// TIA Portal project "Label_Process" (V20)
// Label and sorter box process

(* hardware
DEVICE "S7-1200 station_1"  S7-1200 Station
   slot 0: "Rack_0"  S7-1200 Rack  Rack  V1.0
   slot 1: "PLC_1"  CPU 1212C AC/DC/Rly  6ES7 212-1BE40-0XB0  V4.6
DEVICE "HMI_1"  TP1200 Comfort
   slot 0: "HMI_1"  TP1200 Comfort  6AV2 124-0MC01-0AX0  17.0.0.0
   slot 1: "HMI_RT_1"  TP1200 Comfort  6AV2 124-0MC01-0AX0  17.0.0.0
   slot 5: "HMI_1.IE_CP_1"  PROFINET Interface  17.0.0.0
      slot 1: "PROFINET Interface_1"  PROFINET Interface
         slot 1: "Port_1"  Port
         slot 2: "Port_2"  Port
   slot 7: "HMI_1.MPI/DP_CP_1"  MPI/DP Interface  17.0.0.0
*)

// ===== PLC "PLC_1"  CPU 1212C AC/DC/Rly =====

VAR_GLOBAL   // PLC tag table "Inputs_FactoryIO"
   "Emergency_Stop" AT %I1.0 : Bool;   // Emergency stop mushroom
   "Stop_Pb" AT %I1.1 : Bool;   // Stop pushbutton
   "Start_Pb" AT %I1.2 : Bool;   // Start pushbutton
   "Pause_Signal" AT %I1.3 : Bool;   // Selector for pause process
   "Heigh_Box" AT %I1.4 : Bool;   // Sensor for heigh box
   "Position_Box" AT %I1.5 : Bool;   // Sensor of position box at the label zone
   "Unlabel_Box" AT %I1.6 : Bool;   // Unlabel box sensor
   "Thermal_Fault" AT %I1.7 : Bool;   // Thermal Fault from thermal relays
   "Clock_Byte" AT %MB10 : Byte;
   "Clock_10Hz" AT %M10.0 : Bool;
   "Clock_5Hz" AT %M10.1 : Bool;
   "Clock_2.5Hz" AT %M10.2 : Bool;
   "Clock_2Hz" AT %M10.3 : Bool;
   "Clock_1.25Hz" AT %M10.4 : Bool;
   "Clock_1Hz" AT %M10.5 : Bool;
   "Clock_0.625Hz" AT %M10.6 : Bool;
   "Clock_0.5Hz" AT %M10.7 : Bool;
   "Tag_1" AT %M8.1 : Bool;
   "Tag_2" AT %M1.1 : Bool;
END_VAR

VAR_GLOBAL   // PLC tag table "Outputs"
   "Conveyor M1" AT %Q0.0 : Bool;   // Control Conveyor Belt M1
   "Conveyor M2" AT %Q0.1 : Bool;   // Control Conveyor Belt M2
   "Conveyor M3" AT %Q0.2 : Bool;   // Control Conveyor Belt M3
   "Sorter" AT %Q0.3 : Bool;   // Activate sorter
   "Sorter_Left" AT %Q0.4 : Bool;   // Activate sorter for left position
   "Axis_Label" AT %Q0.5 : Bool;   // Axis control for labeled
END_VAR

DATA_BLOCK "DATA"   // DB1
{ S7_Optimized_Access := 'TRUE' }
VERSION : 0.1
   VAR
      varCounters : Struct
         Labeled_Boxes_Counter : Int;   // Labeled boxes counter
         Unlabel_Boxes_Counter : Int;   // Unlabel boxes counter
         CountUp_Unlabel : Bool;
         Total_Boxes : Int;
         Reset_Counters : Bool;
         Label_TimeSec : DInt;
      END_STRUCT;
      activateSorter : Struct
         M_Sorter_Left : Bool;
         M1_Activate_Sorter : Bool;
         M2_Activate_Sorter : Bool;
      END_STRUCT;
      risingEgde : Struct
         R_StartPB : Bool;   // Memory for rising edge Start button
         R_positionBox : Bool;   // Memory for rising edge position box sensor
         R_Heigh_Box : Bool;   // Memory for rising egde heigh box sensor
         R_Unlabel_Box : Bool;   // Memory for rising egde unlabel box sensor
         R_CountUP_Unlabel : Bool;
         R_Move_CountUP : Bool;
      END_STRUCT;
      generalData : Struct
         M_startStop : Bool;   // Memory for Start Stop all process
         M_pauseProcess : Bool;   // Memory for Pause all process
      END_STRUCT;
      Belts_Data : Struct
         M_Activate_M1 : Bool;   // Memory for activate Belt Conveyor M1
         M_Activate_M2 : Bool;   // Memory for activate Belt Conveyor M2
         M_Activate_M3 : Bool;   // Memory for activate Belt Conveyor M3
      END_STRUCT;
   END_VAR
BEGIN
END_DATA_BLOCK

DATA_BLOCK "HMI_Data"   // DB3
{ S7_Optimized_Access := 'TRUE' }
VERSION : 0.1
   VAR
      "Inputs from HMI" : Struct   // Inputs signals from HMI
         startSignal : Bool;   // Start all process
         stopSignal : Bool;   // Stop all process
         resetCounters : Bool;   // Reset all counters
         pauseProcess : Bool;   // Pause all process
      END_STRUCT;
      Move_Animation : Int;   // HMI box animation
      "Belt Control" : Struct   // Start signals for each belt conveyor
         Start_M1 : Bool;   // Start belt conveyor M1
         Start_M2 : Bool;   // Start belt conveyor M2
         Start_M3 : Bool;   // Start belt conveyor M3
      END_STRUCT;
      "Sorter & Axis Control" : Struct   // Controlling sorter and axis label
         activateAxis : Bool;
         activateSorter : Bool;
         activateSorterLeft : Bool;
      END_STRUCT;
      Counters : Struct
         resetCounterLabeled : Bool;
         resetCounterUnlabel : Bool;
         labelTime : DInt;
      END_STRUCT;
   END_VAR
BEGIN
END_DATA_BLOCK

DATA_BLOCK "HMI_Alarms"   // DB4
{ S7_Optimized_Access := 'FALSE' }
VERSION : 0.1
   VAR
      noTimeSet : Bool;   // Alarm indicator, no time for axis label actuator
      emergencyStopPushed : Bool;   // Alarm indicator, emergency stop pushed
      thermalFault : Bool;   // Alarm indicator, fault thermal relays
      pauseActive : Bool;   // Warning indicator, pause active
   END_VAR
BEGIN
END_DATA_BLOCK

// folder: System blocks/Program resources

DATA_BLOCK "axisTimer"   // DB2
{ S7_Optimized_Access := 'TRUE' }
AUTHOR : Simatic
FAMILY : IEC
NAME : IEC_TMR
VERSION : 1.0
// stored: InstanceOfName IEC_TIMER
"IEC_TIMER"
BEGIN
END_DATA_BLOCK

// folder: (top level)

FUNCTION "Start_Stop" : Void   // FC1, LAD
TITLE = Start and Stop Block
{ S7_Optimized_Access := 'TRUE' }
AUTHOR : Stiven Perez
VERSION : 0.1
// Start and stop conditions to all process
   VAR_INPUT
      emergencyStop : Bool;   // Emergency stop mushroom
      stopPB : Bool;   // Stop Pushbutton
      startPB : Bool;   // Start Pushbutton
      pauseSignal : Bool;   // Pause Selector signal
      HMI_Start : Bool;
      HMI_Stop : Bool;
      HMI_Pause : Bool;
      HMI_Reset_CounterLabel : Bool;
      HMI_Reset_CounterUnlabel : Bool;
      thermalFault : Bool;   // Thermal Fault from thermal relays
   END_VAR
   VAR_OUTPUT
      M_Pause : Bool;   // Memory for Pause process
      emergencyStopAlarm : Bool;
      noTimeSetAlarm : Bool;
      thermalFaultAlarm : Bool;
      pauseActiveWarning : Bool;
      pau : Int;
   END_VAR
   VAR_IN_OUT
      M_startStop : Bool;   // Memory for Start Stop
      labeledCounter : Int;
      unlabelCounter : Int;
      resetCounters : Bool;
   END_VAR
   VAR_TEMP   // added for the SCL form of the ladder/FBD networks
      _w1 : Bool;
   END_VAR
BEGIN

REGION Network 1: Memory for Start Stop
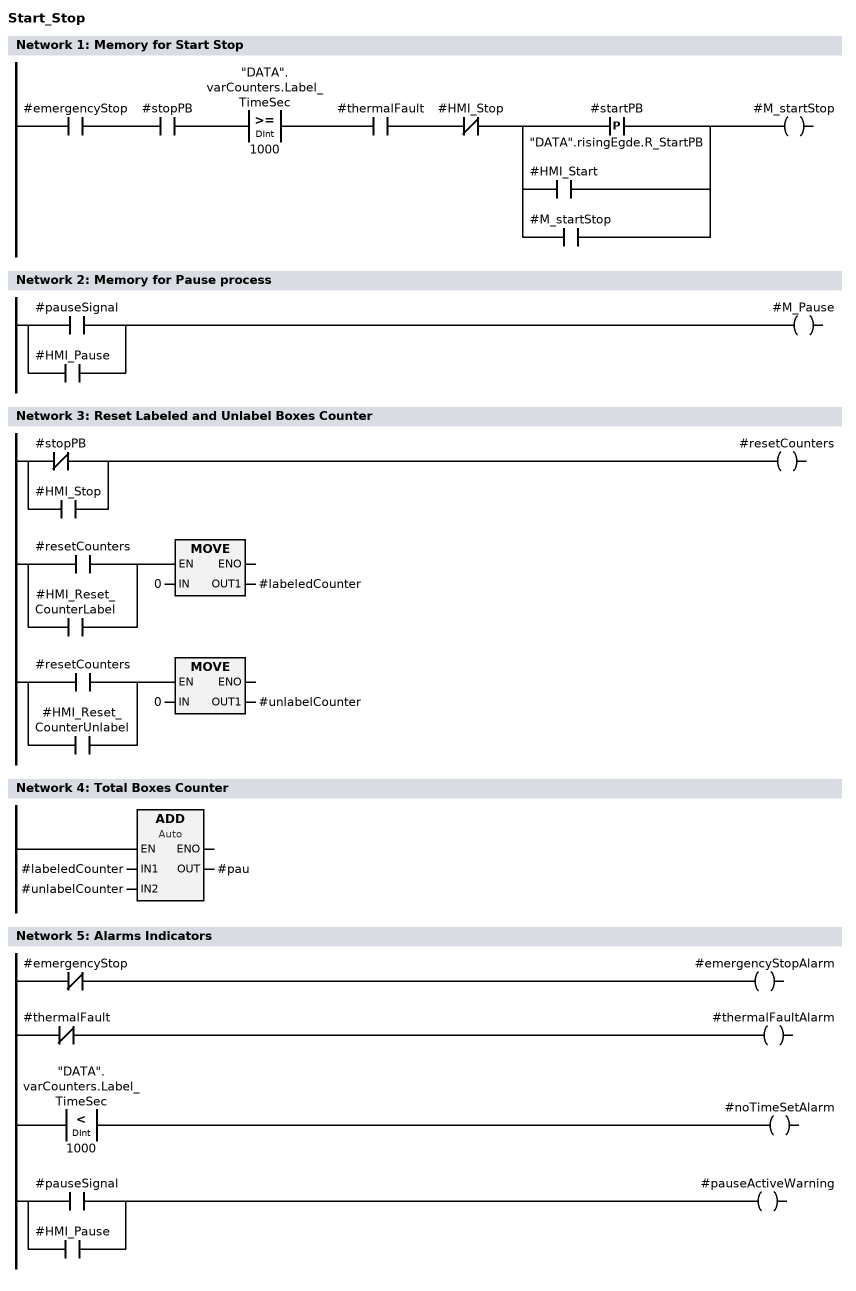
   RUNG wire#powerrail
      Contact( #emergencyStop )
      Contact( #stopPB )
      { S7_Templates := "SrcType := DInt" } GE_Contact(in1 := "DATA".varCounters.Label_TimeSec, in2 := 1000)
      Contact( #thermalFault )
      I_Contact( #HMI_Stop )
      wire#w1
      P_Contact(operand := #startPB, bit := "DATA".risingEgde.R_StartPB)
      wire#w2
      Coil( #M_startStop )
   END_RUNG
   RUNG wire#w1
      Contact( #HMI_Start )
   END_RUNG wire#w2
   RUNG wire#w1
      Contact( #M_startStop )
   END_RUNG wire#w2
   // the same network as SCL:
   #_w1 := #emergencyStop AND #stopPB AND ("DATA".varCounters.Label_TimeSec >= 1000) AND #thermalFault AND NOT #HMI_Stop AND #startPB AND NOT "DATA".risingEgde.R_StartPB;   // rising edge of #startPB
   "DATA".risingEgde.R_StartPB := #startPB;
   #M_startStop := #_w1 OR (#emergencyStop AND #stopPB AND ("DATA".varCounters.Label_TimeSec >= 1000) AND #thermalFault AND NOT #HMI_Stop AND (#HMI_Start OR #M_startStop));
END_REGION

REGION Network 2: Memory for Pause process
   RUNG wire#powerrail
      Contact( #pauseSignal )
      wire#w1
      Coil( #M_Pause )
   END_RUNG
   RUNG wire#powerrail
      Contact( #HMI_Pause )
   END_RUNG wire#w1
   // the same network as SCL:
   #M_Pause := #pauseSignal OR #HMI_Pause;
END_REGION

REGION Network 3: Reset Labeled and Unlabel Boxes Counter
   RUNG wire#powerrail
      I_Contact( #stopPB )
      wire#w1
      Coil( #resetCounters )
   END_RUNG
   RUNG wire#powerrail
      Contact( #HMI_Stop )
   END_RUNG wire#w1
   RUNG wire#powerrail
      Contact( #resetCounters )
      wire#w2
      Move(in := 0, out1 => #labeledCounter)
   END_RUNG
   RUNG wire#powerrail
      Contact( #HMI_Reset_CounterLabel )
   END_RUNG wire#w2
   RUNG wire#powerrail
      Contact( #resetCounters )
      wire#w3
      Move(in := 0, out1 => #unlabelCounter)
   END_RUNG
   RUNG wire#powerrail
      Contact( #HMI_Reset_CounterUnlabel )
   END_RUNG wire#w3
   // the same network as SCL:
   #resetCounters := NOT #stopPB OR #HMI_Stop;
   IF #resetCounters OR #HMI_Reset_CounterLabel THEN #labeledCounter := 0; END_IF;
   IF #resetCounters OR #HMI_Reset_CounterUnlabel THEN #unlabelCounter := 0; END_IF;
END_REGION

REGION Network 4: Total Boxes Counter
   RUNG wire#powerrail
      Add(in1 := #labeledCounter, in2 := #unlabelCounter, out => #pau)
   END_RUNG
   // the same network as SCL:
   #pau := #labeledCounter + #unlabelCounter;
END_REGION

REGION Network 5: Alarms Indicators
   RUNG wire#powerrail
      I_Contact( #emergencyStop )
      Coil( #emergencyStopAlarm )
   END_RUNG
   RUNG wire#powerrail
      I_Contact( #thermalFault )
      Coil( #thermalFaultAlarm )
   END_RUNG
   RUNG wire#powerrail
      { S7_Templates := "SrcType := DInt" } LT_Contact(in1 := "DATA".varCounters.Label_TimeSec, in2 := 1000)
      Coil( #noTimeSetAlarm )
   END_RUNG
   RUNG wire#powerrail
      Contact( #pauseSignal )
      wire#w1
      Coil( #pauseActiveWarning )
   END_RUNG
   RUNG wire#powerrail
      Contact( #HMI_Pause )
   END_RUNG wire#w1
   // the same network as SCL:
   #emergencyStopAlarm := NOT #emergencyStop;
   #thermalFaultAlarm := NOT #thermalFault;
   #noTimeSetAlarm := "DATA".varCounters.Label_TimeSec < 1000;
   #pauseActiveWarning := #pauseSignal OR #HMI_Pause;
END_REGION
END_FUNCTION

FUNCTION "Box_Labeling" : Void   // FC2, LAD
TITLE = Box Sorting Block
{ S7_Optimized_Access := 'TRUE' }
AUTHOR : Stiven Perez
VERSION : 0.1
// Conditions to select the correct box to labeled
   VAR_INPUT
      M_startStop : Bool;
      M_pauseSignal : Bool;
      positionBox : Bool;
      HMI_Start_M1 : Bool;
      HMI_Start_M2 : Bool;
      Label_Time : DInt;
      HMI_Activate_Axis : Bool;
   END_VAR
   VAR_OUTPUT
      conveyorM1 : Bool;   // Conveyor M1 Start
      conveyorM2 : Bool;   // Conveyor M2 Start
      M1_activateSorter : Bool;   // Memory for activate sorter
   END_VAR
   VAR_IN_OUT
      axisControl : Bool;
      labeledBoxes_Counter : Int;
      M_Activate_M1 : Bool;   // Memory for activate Belt M1
      M_Activate_M2 : Bool;   // Memory for activate Belt M2
      Label_Time_Sec : DInt;
   END_VAR
   VAR_TEMP   // added for the SCL form of the ladder/FBD networks
      _w1 : Bool;
      _w2 : Bool;
   END_VAR
BEGIN

REGION Network 1: Activate Conveyor Belts 1, 2 and Sorter
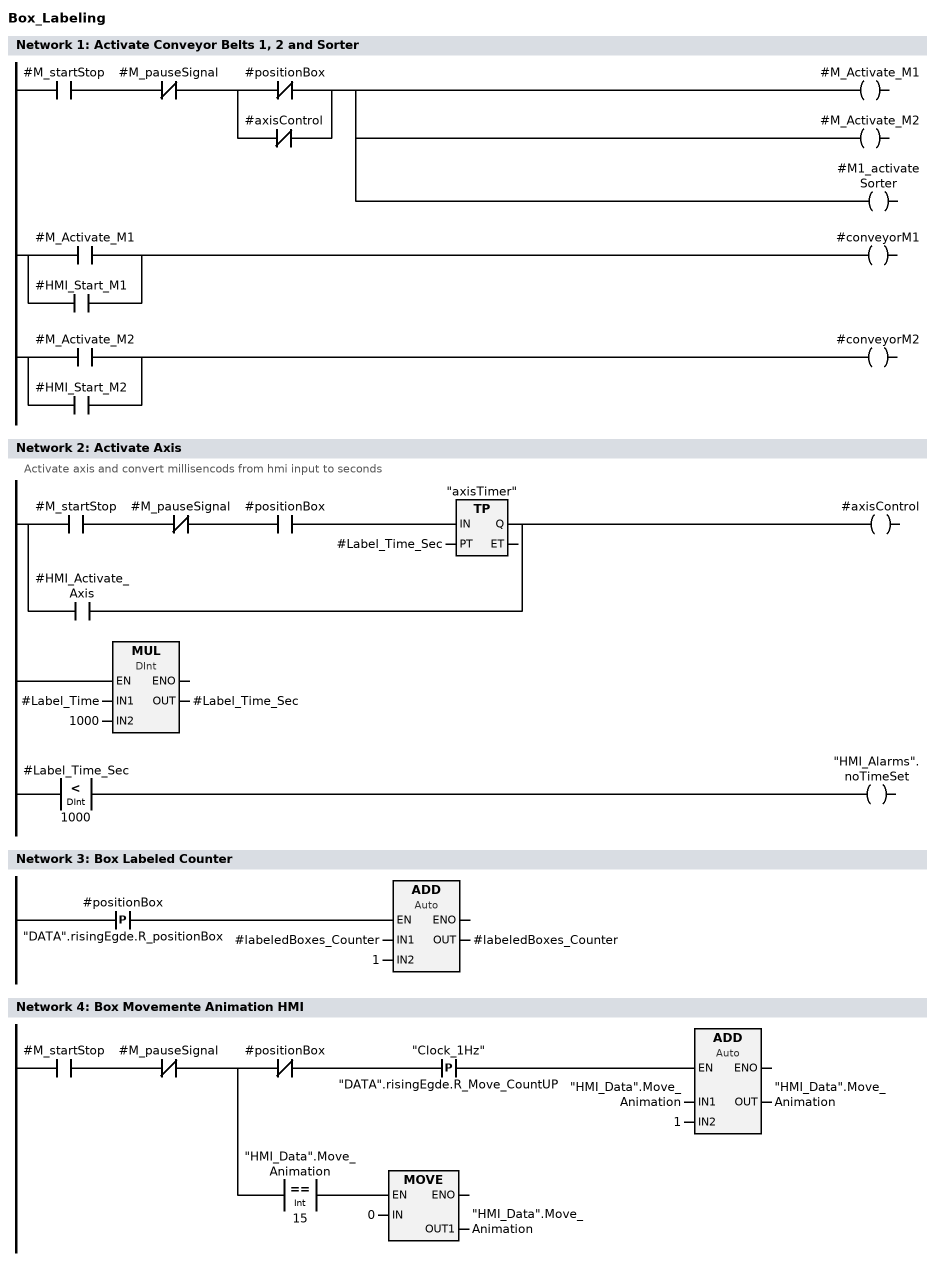
   RUNG wire#powerrail
      Contact( #M_startStop )
      I_Contact( #M_pauseSignal )
      wire#w1
      I_Contact( #positionBox )
      wire#w2
      Coil( #M_Activate_M1 )
   END_RUNG
   RUNG wire#w1
      I_Contact( #axisControl )
   END_RUNG wire#w2
   RUNG wire#w2
      Coil( #M_Activate_M2 )
   END_RUNG
   RUNG wire#w2
      Coil( #M1_activateSorter )
   END_RUNG
   RUNG wire#powerrail
      Contact( #M_Activate_M1 )
      wire#w3
      Coil( #conveyorM1 )
   END_RUNG
   RUNG wire#powerrail
      Contact( #HMI_Start_M1 )
   END_RUNG wire#w3
   RUNG wire#powerrail
      Contact( #M_Activate_M2 )
      wire#w4
      Coil( #conveyorM2 )
   END_RUNG
   RUNG wire#powerrail
      Contact( #HMI_Start_M2 )
   END_RUNG wire#w4
   // the same network as SCL:
   #M_Activate_M1 := #M_startStop AND NOT #M_pauseSignal AND (NOT #positionBox OR NOT #axisControl);
   #M_Activate_M2 := #M_Activate_M1;
   #M1_activateSorter := #M_Activate_M1;
   #conveyorM1 := #M_Activate_M1 OR #HMI_Start_M1;
   #conveyorM2 := #M_Activate_M2 OR #HMI_Start_M2;
END_REGION

REGION Network 2: Activate Axis
   // Activate axis and convert millisencods from hmi input to seconds
   "axisTimer".TP(IN := #M_startStop AND NOT #M_pauseSignal AND #positionBox, PT := #Label_Time_Sec);
   #axisControl := "axisTimer".Q OR #HMI_Activate_Axis;
   #Label_Time_Sec := #Label_Time * 1000;
   "HMI_Alarms".noTimeSet := #Label_Time_Sec < 1000;
END_REGION

REGION Network 3: Box Labeled Counter
   RUNG wire#powerrail
      P_Contact(operand := #positionBox, bit := "DATA".risingEgde.R_positionBox)
      Add(in1 := #labeledBoxes_Counter, in2 := 1, out => #labeledBoxes_Counter)
   END_RUNG
   // the same network as SCL:
   #_w1 := #positionBox AND NOT "DATA".risingEgde.R_positionBox;   // rising edge of #positionBox
   "DATA".risingEgde.R_positionBox := #positionBox;
   IF #_w1 THEN #labeledBoxes_Counter := #labeledBoxes_Counter + 1; END_IF;
END_REGION

REGION Network 4: Box Movemente Animation HMI
   RUNG wire#powerrail
      Contact( #M_startStop )
      I_Contact( #M_pauseSignal )
      wire#w1
      I_Contact( #positionBox )
      P_Contact(operand := "Clock_1Hz", bit := "DATA".risingEgde.R_Move_CountUP)
      Add(in1 := "HMI_Data".Move_Animation, in2 := 1, out => "HMI_Data".Move_Animation)
   END_RUNG
   RUNG wire#w1
      { S7_Templates := "SrcType := Int" } EQ_Contact(in1 := "HMI_Data".Move_Animation, in2 := 15)
      Move(in := 0, out1 => "HMI_Data".Move_Animation)
   END_RUNG
   // the same network as SCL:
   #_w1 := #M_startStop AND NOT #M_pauseSignal;
   #_w2 := #_w1 AND NOT #positionBox AND "Clock_1Hz" AND NOT "DATA".risingEgde.R_Move_CountUP;   // rising edge of "Clock_1Hz"
   "DATA".risingEgde.R_Move_CountUP := "Clock_1Hz";
   IF #_w2 THEN "HMI_Data".Move_Animation := "HMI_Data".Move_Animation + 1; END_IF;
   IF #_w1 AND ("HMI_Data".Move_Animation = 15) THEN "HMI_Data".Move_Animation := 0; END_IF;
END_REGION
END_FUNCTION

FUNCTION "Unlabeled_Boxes" : Void   // FC3, LAD
TITLE = Unlabeled Boxes Block
{ S7_Optimized_Access := 'TRUE' }
AUTHOR : Stiven Perez
VERSION : 0.1
// Conditions to activate left sorter and unlabeled counter, this function will be activate when the heigh box is out of range
   VAR_INPUT
      M_startStop : Bool;
      M_pauseSignal : Bool;
      heighBox : Bool;
      Unlabel_Box : Bool;
      HMI_Start_M3 : Bool;
      HMI_Activate_SorterLeft : Bool;
      HMI_Activate_Sorter : Bool;
   END_VAR
   VAR_OUTPUT
      conveyorM3 : Bool;
      sorterLeft : Bool;
      sorter : Bool;
   END_VAR
   VAR_IN_OUT
      M1_activateSorter : Bool;
      M2_activateSorter : Bool;
      countUp_Unlabel : Bool;
      unlabelBoxes_Counter : Int;
   END_VAR
   VAR_TEMP   // added for the SCL form of the ladder/FBD networks
      _w1 : Bool;
      _w2 : Bool;
      _w3 : Bool;
   END_VAR
BEGIN

REGION Network 1: Activate Belt Conveyor 3
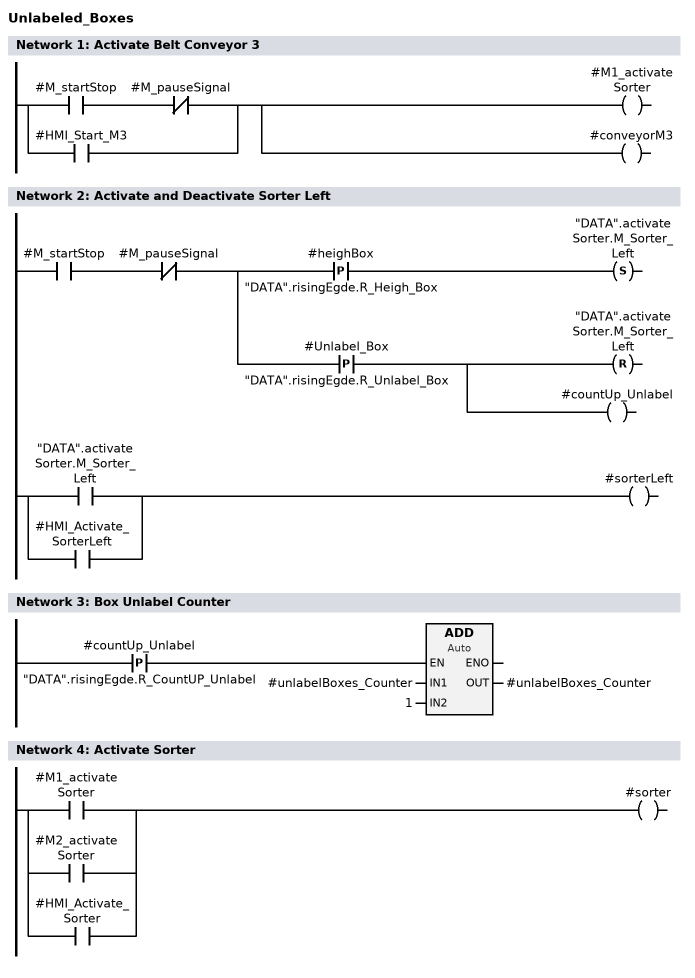
   RUNG wire#powerrail
      Contact( #M_startStop )
      I_Contact( #M_pauseSignal )
      wire#w1
      Coil( #M1_activateSorter )
   END_RUNG
   RUNG wire#powerrail
      Contact( #HMI_Start_M3 )
   END_RUNG wire#w1
   RUNG wire#w1
      Coil( #conveyorM3 )
   END_RUNG
   // the same network as SCL:
   #M1_activateSorter := (#M_startStop AND NOT #M_pauseSignal) OR #HMI_Start_M3;
   #conveyorM3 := #M1_activateSorter;
END_REGION

REGION Network 2: Activate and Deactivate Sorter Left
   RUNG wire#powerrail
      Contact( #M_startStop )
      I_Contact( #M_pauseSignal )
      wire#w1
      P_Contact(operand := #heighBox, bit := "DATA".risingEgde.R_Heigh_Box)
      S_Coil( "DATA".activateSorter.M_Sorter_Left )
   END_RUNG
   RUNG wire#w1
      P_Contact(operand := #Unlabel_Box, bit := "DATA".risingEgde.R_Unlabel_Box)
      wire#w2
      R_Coil( "DATA".activateSorter.M_Sorter_Left )
   END_RUNG
   RUNG wire#w2
      Coil( #countUp_Unlabel )
   END_RUNG
   RUNG wire#powerrail
      Contact( "DATA".activateSorter.M_Sorter_Left )
      wire#w3
      Coil( #sorterLeft )
   END_RUNG
   RUNG wire#powerrail
      Contact( #HMI_Activate_SorterLeft )
   END_RUNG wire#w3
   // the same network as SCL:
   #_w1 := #M_startStop AND NOT #M_pauseSignal;
   #_w2 := #_w1 AND #heighBox AND NOT "DATA".risingEgde.R_Heigh_Box;   // rising edge of #heighBox
   "DATA".risingEgde.R_Heigh_Box := #heighBox;
   IF #_w2 THEN "DATA".activateSorter.M_Sorter_Left := TRUE; END_IF;
   #_w3 := #_w1 AND #Unlabel_Box AND NOT "DATA".risingEgde.R_Unlabel_Box;   // rising edge of #Unlabel_Box
   "DATA".risingEgde.R_Unlabel_Box := #Unlabel_Box;
   IF #_w3 THEN "DATA".activateSorter.M_Sorter_Left := FALSE; END_IF;
   #countUp_Unlabel := #_w3;
   #sorterLeft := "DATA".activateSorter.M_Sorter_Left OR #HMI_Activate_SorterLeft;
END_REGION

REGION Network 3: Box Unlabel Counter
   RUNG wire#powerrail
      P_Contact(operand := #countUp_Unlabel, bit := "DATA".risingEgde.R_CountUP_Unlabel)
      Add(in1 := #unlabelBoxes_Counter, in2 := 1, out => #unlabelBoxes_Counter)
   END_RUNG
   // the same network as SCL:
   #_w1 := #countUp_Unlabel AND NOT "DATA".risingEgde.R_CountUP_Unlabel;   // rising edge of #countUp_Unlabel
   "DATA".risingEgde.R_CountUP_Unlabel := #countUp_Unlabel;
   IF #_w1 THEN #unlabelBoxes_Counter := #unlabelBoxes_Counter + 1; END_IF;
END_REGION

REGION Network 4: Activate Sorter
   RUNG wire#powerrail
      Contact( #M1_activateSorter )
      wire#w1
      Coil( #sorter )
   END_RUNG
   RUNG wire#powerrail
      Contact( #M2_activateSorter )
   END_RUNG wire#w1
   RUNG wire#powerrail
      Contact( #HMI_Activate_Sorter )
   END_RUNG wire#w1
   // the same network as SCL:
   #sorter := #M1_activateSorter OR #M2_activateSorter OR #HMI_Activate_Sorter;
END_REGION
END_FUNCTION

ORGANIZATION_BLOCK "Main"   // OB1, LAD, ProgramCycle
TITLE = "Main Program Sweep (Cycle)"
{ S7_Optimized_Access := 'TRUE' }
VERSION : 0.1
   VAR_INPUT
      Initial_Call : Bool;   // Initial call of this OB
      Remanence : Bool;   // =True, if remanent data are available
   END_VAR
BEGIN

REGION Network 1: Start-stop for all process
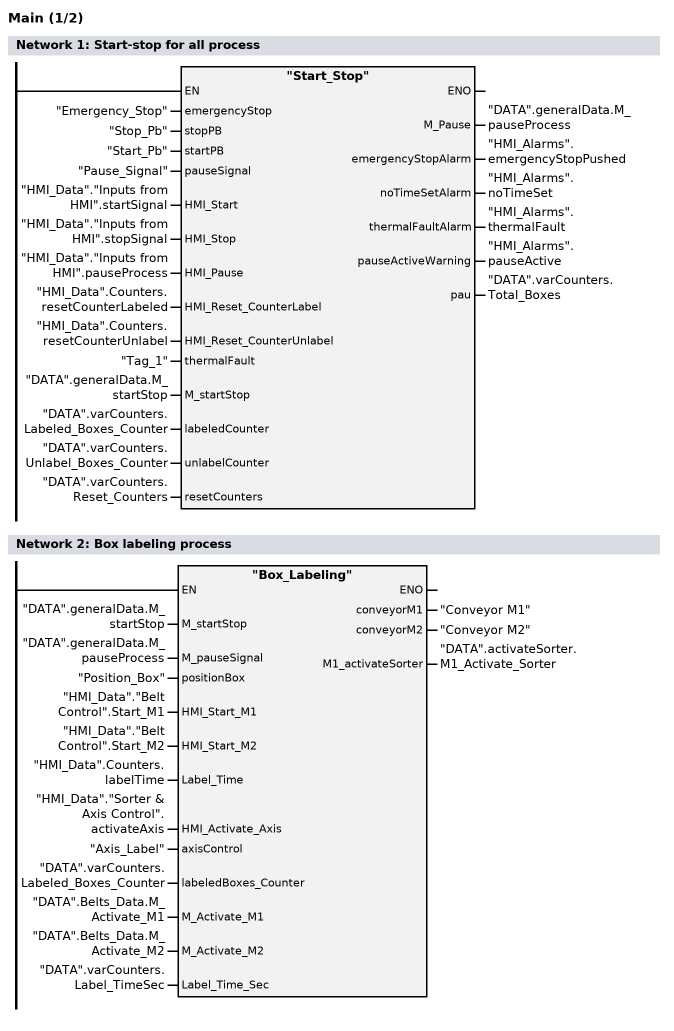
   RUNG wire#powerrail
      "Start_Stop"(emergencyStop := "Emergency_Stop", stopPB := "Stop_Pb", startPB := "Start_Pb", pauseSignal := "Pause_Signal", HMI_Start := "HMI_Data"."Inputs from HMI".startSignal, HMI_Stop := "HMI_Data"."Inputs from HMI".stopSignal, HMI_Pause := "HMI_Data"."Inputs from HMI".pauseProcess, HMI_Reset_CounterLabel := "HMI_Data".Counters.resetCounterLabeled, HMI_Reset_CounterUnlabel := "HMI_Data".Counters.resetCounterUnlabel, thermalFault := "Tag_1", M_startStop := "DATA".generalData.M_startStop, labeledCounter := "DATA".varCounters.Labeled_Boxes_Counter, unlabelCounter := "DATA".varCounters.Unlabel_Boxes_Counter, resetCounters := "DATA".varCounters.Reset_Counters, M_Pause => "DATA".generalData.M_pauseProcess, emergencyStopAlarm => "HMI_Alarms".emergencyStopPushed, noTimeSetAlarm => "HMI_Alarms".noTimeSet, thermalFaultAlarm => "HMI_Alarms".thermalFault, pauseActiveWarning => "HMI_Alarms".pauseActive, pau => "DATA".varCounters.Total_Boxes)
   END_RUNG
   // the same network as SCL:
   "Start_Stop"(emergencyStop := "Emergency_Stop",
                stopPB := "Stop_Pb",
                startPB := "Start_Pb",
                pauseSignal := "Pause_Signal",
                HMI_Start := "HMI_Data"."Inputs from HMI".startSignal,
                HMI_Stop := "HMI_Data"."Inputs from HMI".stopSignal,
                HMI_Pause := "HMI_Data"."Inputs from HMI".pauseProcess,
                HMI_Reset_CounterLabel := "HMI_Data".Counters.resetCounterLabeled,
                HMI_Reset_CounterUnlabel := "HMI_Data".Counters.resetCounterUnlabel,
                thermalFault := "Tag_1",
                M_startStop := "DATA".generalData.M_startStop,
                labeledCounter := "DATA".varCounters.Labeled_Boxes_Counter,
                unlabelCounter := "DATA".varCounters.Unlabel_Boxes_Counter,
                resetCounters := "DATA".varCounters.Reset_Counters,
                M_Pause => "DATA".generalData.M_pauseProcess,
                emergencyStopAlarm => "HMI_Alarms".emergencyStopPushed,
                noTimeSetAlarm => "HMI_Alarms".noTimeSet,
                thermalFaultAlarm => "HMI_Alarms".thermalFault,
                pauseActiveWarning => "HMI_Alarms".pauseActive,
                pau => "DATA".varCounters.Total_Boxes);
END_REGION

REGION Network 2: Box labeling process
   RUNG wire#powerrail
      "Box_Labeling"(M_startStop := "DATA".generalData.M_startStop, M_pauseSignal := "DATA".generalData.M_pauseProcess, positionBox := "Position_Box", HMI_Start_M1 := "HMI_Data"."Belt Control".Start_M1, HMI_Start_M2 := "HMI_Data"."Belt Control".Start_M2, Label_Time := "HMI_Data".Counters.labelTime, HMI_Activate_Axis := "HMI_Data"."Sorter & Axis Control".activateAxis, axisControl := "Axis_Label", labeledBoxes_Counter := "DATA".varCounters.Labeled_Boxes_Counter, M_Activate_M1 := "DATA".Belts_Data.M_Activate_M1, M_Activate_M2 := "DATA".Belts_Data.M_Activate_M2, Label_Time_Sec := "DATA".varCounters.Label_TimeSec, conveyorM1 => "Conveyor M1", conveyorM2 => "Conveyor M2", M1_activateSorter => "DATA".activateSorter.M1_Activate_Sorter)
   END_RUNG
   // the same network as SCL:
   "Box_Labeling"(M_startStop := "DATA".generalData.M_startStop,
                  M_pauseSignal := "DATA".generalData.M_pauseProcess,
                  positionBox := "Position_Box",
                  HMI_Start_M1 := "HMI_Data"."Belt Control".Start_M1,
                  HMI_Start_M2 := "HMI_Data"."Belt Control".Start_M2,
                  Label_Time := "HMI_Data".Counters.labelTime,
                  HMI_Activate_Axis := "HMI_Data"."Sorter & Axis Control".activateAxis,
                  axisControl := "Axis_Label",
                  labeledBoxes_Counter := "DATA".varCounters.Labeled_Boxes_Counter,
                  M_Activate_M1 := "DATA".Belts_Data.M_Activate_M1,
                  M_Activate_M2 := "DATA".Belts_Data.M_Activate_M2,
                  Label_Time_Sec := "DATA".varCounters.Label_TimeSec,
                  conveyorM1 => "Conveyor M1",
                  conveyorM2 => "Conveyor M2",
                  M1_activateSorter => "DATA".activateSorter.M1_Activate_Sorter);
END_REGION

REGION Network 3: Unlabeled boxes process
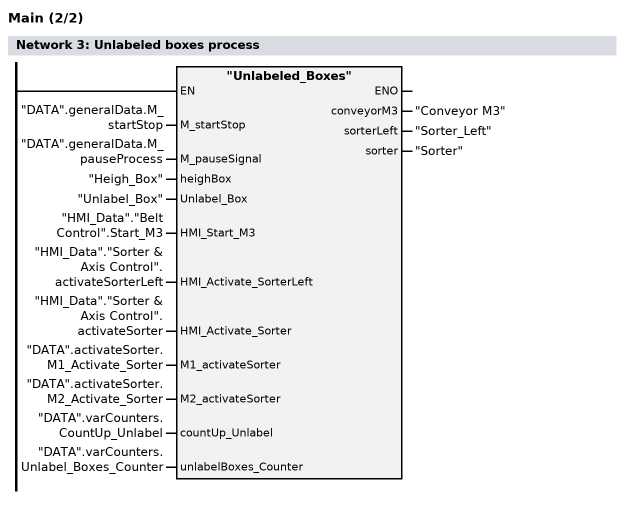
   RUNG wire#powerrail
      "Unlabeled_Boxes"(M_startStop := "DATA".generalData.M_startStop, M_pauseSignal := "DATA".generalData.M_pauseProcess, heighBox := "Heigh_Box", Unlabel_Box := "Unlabel_Box", HMI_Start_M3 := "HMI_Data"."Belt Control".Start_M3, HMI_Activate_SorterLeft := "HMI_Data"."Sorter & Axis Control".activateSorterLeft, HMI_Activate_Sorter := "HMI_Data"."Sorter & Axis Control".activateSorter, M1_activateSorter := "DATA".activateSorter.M1_Activate_Sorter, M2_activateSorter := "DATA".activateSorter.M2_Activate_Sorter, countUp_Unlabel := "DATA".varCounters.CountUp_Unlabel, unlabelBoxes_Counter := "DATA".varCounters.Unlabel_Boxes_Counter, conveyorM3 => "Conveyor M3", sorterLeft => "Sorter_Left", sorter => "Sorter")
   END_RUNG
   // the same network as SCL:
   "Unlabeled_Boxes"(M_startStop := "DATA".generalData.M_startStop,
                     M_pauseSignal := "DATA".generalData.M_pauseProcess,
                     heighBox := "Heigh_Box",
                     Unlabel_Box := "Unlabel_Box",
                     HMI_Start_M3 := "HMI_Data"."Belt Control".Start_M3,
                     HMI_Activate_SorterLeft := "HMI_Data"."Sorter & Axis Control".activateSorterLeft,
                     HMI_Activate_Sorter := "HMI_Data"."Sorter & Axis Control".activateSorter,
                     M1_activateSorter := "DATA".activateSorter.M1_Activate_Sorter,
                     M2_activateSorter := "DATA".activateSorter.M2_Activate_Sorter,
                     countUp_Unlabel := "DATA".varCounters.CountUp_Unlabel,
                     unlabelBoxes_Counter := "DATA".varCounters.Unlabel_Boxes_Counter,
                     conveyorM3 => "Conveyor M3",
                     sorterLeft => "Sorter_Left",
                     sorter => "Sorter");
END_REGION
END_ORGANIZATION_BLOCK

(* ===== HMI "HMI_RT_1" =====
system functions are stored by id; their names below are inferred from use
connection "HMI_Connection_1": ETHERNET, S7_1200_OMS

HMI tags "Actuators"
   "axisLabel" : Bool = PLC Axis_Label AT %Q0.5, 1 s   // Run signal indicator
   "conveyor_M3" : Bool = PLC "Conveyor M3" AT %Q0.2, 1 s   // Run signal indicator
   "conveyor_M2" : Bool = PLC "Conveyor M2" AT %Q0.1, 1 s   // Run signal indicator
   "conveyor_M1" : Bool = PLC "Conveyor M1" AT %Q0.0, 1 s   // Run signal indicator
   "unlabelBox" : Bool = PLC Unlabel_Box AT %I1.6, 100 ms   // Activate signal indicator
   "heighBox" : Bool = PLC Heigh_Box AT %I1.4, 100 ms   // Activate signal indicator
   "positionBox" : Bool = PLC Position_Box AT %I1.5, 100 ms   // Activate signal indicator
   "sorter" : Bool = PLC Sorter AT %Q0.3, 1 s
   "sorterLeft" : Bool = PLC Sorter_Left AT %Q0.4, 1 s

HMI tags "Inputs"
   "startSignal" : Bool = PLC HMI_Data."Inputs from HMI".startSignal AT %DB1.DBX0.0, 1 s
   "stopSignal" : Bool = PLC HMI_Data."Inputs from HMI".stopSignal AT %DB1.DBX0.0, 1 s
   "pauseProcess" : Bool = PLC HMI_Data."Inputs from HMI".pauseProcess AT %DB1.DBX0.0, 1 s
   "resetCounters" : Bool = PLC HMI_Data."Inputs from HMI".resetCounters AT %DB1.DBX0.0, 1 s
   "thermalFault" : Bool = PLC Tag_1 AT %M8.1, 1 s
   "activateAxis" : Bool = PLC HMI_Data."Sorter & Axis Control".activateAxis AT %DB1.DBX0.0, 1 s
   "activateSorter" : Bool = PLC HMI_Data."Sorter & Axis Control".activateSorter AT %DB1.DBX0.0, 1 s
   "activateSorterLeft" : Bool = PLC HMI_Data."Sorter & Axis Control".activateSorterLeft AT %DB1.DBX0.0, 1 s
   "startM1" : Bool = PLC HMI_Data."Belt Control".Start_M1 AT %DB1.DBX0.0, 1 s
   "startM2" : Bool = PLC HMI_Data."Belt Control".Start_M2 AT %DB1.DBX0.0, 1 s
   "startM3" : Bool = PLC HMI_Data."Belt Control".Start_M3 AT %DB1.DBX0.0, 1 s
   "resetCounterLabeled" : Bool = PLC HMI_Data.Counters.resetCounterLabeled AT %DB1.DBX0.0, 1 s
   "resetCounterUnlabel" : Bool = PLC HMI_Data.Counters.resetCounterUnlabel AT %DB1.DBX0.0, 1 s

HMI tags "Counters"
   "totalCounter" : Int = PLC DATA.varCounters.Total_Boxes AT %DB1.DBW0, 100 ms
   "unlabelBoxesCounter" : Int = PLC DATA.varCounters.Unlabel_Boxes_Counter AT %DB1.DBW0, 100 ms
   "labeledBoxesCounter" : Int = PLC DATA.varCounters.Labeled_Boxes_Counter AT %DB1.DBW0, 100 ms
   "moveAnimation" : Int = PLC HMI_Data.Move_Animation AT %DB1.DBW0, 1 s
   "labelTime" : DInt = PLC HMI_Data.Counters.labelTime AT %DB1.DBW0, 1 s

HMI tags "Global_Vars"
   "startStop" : Bool = PLC DATA.generalData.M_startStop AT %DB1.DBW0, 1 s
   "Tag_ScreenNumber" : Bool AT %DB1.DBX0.0

HMI tags "Alarms"
   "Alarms" : UInt AT %DB4.DBW0, 1 s

discrete alarms
   1: 'No time label set, please enter the label time in Seconds', class Errors, trigger "Alarms" bit 8
   2: 'Emergency Stop has been pushed', class Errors, trigger "Alarms" bit 9
   3: 'Check the thermal relays', class Errors, trigger "Alarms" bit 10
   4: 'The all process in StandBy', class Warnings, trigger "Alarms" bit 11

screen "HomeView" 1280x739, template "Template_1"
   on GenerateScreen: SetTag("Tag_ScreenNumber", 1)
   SymbolLibrary "Symbol library_1" at 315,547 size 838x61
   SymbolLibrary "Symbol library_2" at 457,521 size 105x46
      HorizontalMovement <- "moveAnimation"
      Visibility <- "startStop"
   TextField "Text field_1" at 694,420 size 112x27; Text 'Axis Label'
   SymbolLibrary "Symbol library_3" at 195,62 size 216x107
   SymbolLibrary "Symbol library_5" at 195,62 size 216x107
      Visibility <- "conveyor_M1"
   Circle "Circle_2" at 217,196 size 23x23
      Appearance <- "conveyor_M1"
   Circle "Circle_3" at 217,226 size 23x23
      Appearance <- "conveyor_M1"
   Circle "Circle_4" at 217,256 size 23x23
      Appearance <- "thermalFault"
   TextField "Text field_2" at 274,192 size 42x25; Text 'Run'
   TextField "Text field_3" at 274,222 size 49x25; Text 'Stop'
   TextField "Text field_4" at 273,251 size 53x25; Text 'Fault'
   Circle "Circle_1" at 659,422 size 23x23
      Appearance <- "axisLabel"
   TextField "Text field_5" at 694,452 size 215x27; Text 'Position Box Sensor'
   Circle "Circle_5" at 659,454 size 23x23
      Appearance <- "positionBox"
   IOField "I/O field_1" at 74,388 size 141x57; FormatPattern 9999
      ProcessValue <- "totalCounter"
   TextField "Text field_6" at 78,351 size 139x29; Text 'Total Boxes'
   SymbolLibrary "Symbol library_4" at 544,62 size 216x107
   SymbolLibrary "Symbol library_6" at 544,62 size 216x107
      Visibility <- "conveyor_M2"
   Circle "Circle_6" at 566,196 size 23x23
      Appearance <- "conveyor_M2"
   Circle "Circle_7" at 566,226 size 23x23
      Appearance <- "conveyor_M2"
   Circle "Circle_8" at 566,256 size 23x23
      Appearance <- "thermalFault"
   TextField "Text field_7" at 623,192 size 42x25; Text 'Run'
   TextField "Text field_8" at 623,222 size 49x25; Text 'Stop'
   TextField "Text field_9" at 622,251 size 53x25; Text 'Fault'
   SymbolLibrary "Symbol library_7" at 893,62 size 216x107
   SymbolLibrary "Symbol library_8" at 893,62 size 216x107
      Visibility <- "conveyor_M3"
   Circle "Circle_9" at 915,196 size 23x23
      Appearance <- "conveyor_M3"
   Circle "Circle_10" at 915,226 size 23x23
      Appearance <- "conveyor_M3"
   Circle "Circle_11" at 915,256 size 23x23
      Appearance <- "thermalFault"
   TextField "Text field_10" at 972,192 size 42x25; Text 'Run'
   TextField "Text field_11" at 972,222 size 49x25; Text 'Stop'
   TextField "Text field_12" at 971,251 size 53x25; Text 'Fault'
   TextField "Text field_13" at 192,24 size 190x27; Text 'Belt Conveyor M1'
   TextField "Text field_14" at 543,24 size 190x27; Text 'Belt Conveyor M2'
   TextField "Text field_15" at 892,22 size 190x27; Text 'Belt Conveyor M3'
   IOField "I/O field_2" at 75,491 size 141x57; FormatPattern 9999
      ProcessValue <- "labeledBoxesCounter"
   IOField "I/O field_3" at 76,596 size 141x57; FormatPattern 9999
      ProcessValue <- "unlabelBoxesCounter"
   TextField "Text field_16" at 66,456 size 168x29; Text 'Labeled Boxes'
   TextField "Text field_17" at 70,562 size 166x29; Text 'Unlabel Boxes'

Template "Template_1" 1280x739
   Button "Exit" at 1200,679 size 78x59; TextOff 'Exit'; PictureOff "ExitRuntime_TP1200_Comfort_TR"; PictureOn "ExitRuntime_TP1200_Comfort_TR"
      on Release: StopRuntime(0)
   Button "Template_Button_6" at 917,679 size 78x59; TextOff 'Text'; PictureOff "pausebutton"
      on Press: InvertBit("pauseProcess")
   Button "Template_Button_7" at 813,679 size 78x59; TextOff 'Text'; PictureOff "stop"
      on Press: function_b14e0dd5("stopSignal", 0)
   Button "Template_Button_8" at 710,679 size 78x59; TextOff 'Text'; PictureOff "start-button"
      on Press: function_b14e0dd5("startSignal", 0)
   Button "Template_Button_9" at 571,679 size 78x59; TextOff 'Text'; PictureOff "mechanic"; Authorization "Maintenance"
      on Release: ActivateScreen("Maintenance", 0)
   Button "Template_Button_10" at 422,679 size 78x59; TextOff 'Text'; PictureOff "motor"; Authorization "Maintenance"
      on Release: function_efd93a16("Belt_M3", 400, 125, -1, -1, 1)
   Button "Template_Button_11" at 309,679 size 78x59; TextOff 'Text'; PictureOff "motor"; Authorization "Maintenance"
      on Release: function_efd93a16("Belt_M2", 400, 125, -1, -1, 1)
   Button "Template_Button_12" at 192,678 size 78x59; TextOff 'Text'; PictureOff "motor"; Authorization "Maintenance"
      on Release: function_efd93a16("Belt_M1", 400, 125, -1, -1, 1)
   Button "Alarms" at 1111,679 size 78x59; TextOff 'Alarms'; PictureOff "AlarmDisplay_TP1200_Comfort_TR"; PictureOn "AlarmDisplay_TP1200_Comfort_TR"
      on Release: function_ef3f5d25("System events", -1)
   Button "Start screen" at 1,679 size 78x59; TextOff 'Start screen'; PictureOff "NavigateHome_TP1200_Comfort_TR"; PictureOn "NavigateHome_TP1200_Comfort_TR"
      on Release: ActivateScreen("HomeView", 0)

PopupScreen "Belt_M2" 450x450
   SymbolLibrary "Symbol library_3" at 139,60 size 216x107
   SymbolLibrary "Symbol library_5" at 139,60 size 216x107
      Visibility <- "conveyor_M2"
   Button "Button_1" at 84,235 size 125x61; TextOff 'Start'
      on Release: InvertBit("startM2")
   Circle "Circle_2" at 179,341 size 23x23
      Appearance <- "conveyor_M2"
   Circle "Circle_3" at 179,371 size 23x23
      Appearance <- "conveyor_M2"
   Circle "Circle_4" at 179,401 size 23x23
      Appearance <- "thermalFault"
   TextField "Text field_2" at 232,339 size 42x25; Text 'Run'
   TextField "Text field_3" at 232,369 size 49x25; Text 'Stop'
   TextField "Text field_4" at 232,401 size 53x25; Text 'Fault'
   TextField "Text field_13" at 139,8 size 190x27; Text 'Belt Conveyor M2'
   Button "Button_2" at 268,235 size 125x61; TextOff 'Stop'
      on Release: InvertBit("startM2")

PopupScreen "Belt_M1" 450x450
   SymbolLibrary "Symbol library_3" at 139,60 size 216x107
   SymbolLibrary "Symbol library_5" at 139,60 size 216x107
      Visibility <- "conveyor_M1"
   Button "Button_1" at 84,235 size 125x61; TextOff 'Start'
      on Release: InvertBit("startM1")
   Circle "Circle_2" at 179,341 size 23x23
      Appearance <- "conveyor_M1"
   Circle "Circle_3" at 179,371 size 23x23
      Appearance <- "conveyor_M1"
   Circle "Circle_4" at 179,401 size 23x23
      Appearance <- "thermalFault"
   TextField "Text field_2" at 232,339 size 42x25; Text 'Run'
   TextField "Text field_3" at 232,369 size 49x25; Text 'Stop'
   TextField "Text field_4" at 232,401 size 53x25; Text 'Fault'
   TextField "Text field_13" at 139,8 size 190x27; Text 'Belt Conveyor M1'
   Button "Button_2" at 268,235 size 125x61; TextOff 'Stop'
      on Release: InvertBit("startM1")

PopupScreen "Belt_M3" 450x450
   SymbolLibrary "Symbol library_3" at 139,60 size 216x107
   SymbolLibrary "Symbol library_5" at 139,60 size 216x107
      Visibility <- "conveyor_M3"
   Button "Button_1" at 84,235 size 125x61; TextOff 'Start'
      on Release: InvertBit("startM3")
   Circle "Circle_2" at 179,341 size 23x23
      Appearance <- "conveyor_M3"
   Circle "Circle_3" at 179,371 size 23x23
      Appearance <- "conveyor_M3"
   Circle "Circle_4" at 179,401 size 23x23
      Appearance <- "thermalFault"
   TextField "Text field_2" at 232,339 size 42x25; Text 'Run'
   TextField "Text field_3" at 232,369 size 49x25; Text 'Stop'
   TextField "Text field_4" at 232,401 size 53x25; Text 'Fault'
   TextField "Text field_13" at 139,8 size 190x27; Text 'Belt Conveyor M3'
   Button "Button_2" at 268,235 size 125x61; TextOff 'Stop'
      on Release: InvertBit("startM3")

screen "Maintenance" 1280x739, template "Template_1"
   TextField "Text field_4" at 146,95 size 64x25; Text 'Sorter'
   TextField "Text field_7" at 579,181 size 149x25; Text 'Reset Counters'
   Button "Button_13" at 474,272 size 105x46; TextOff 'Reset'
      on Press: function_b14e0dd5("resetCounterLabeled", 0)
   Button "Button_14" at 694,272 size 105x46; TextOff 'Reset'
      on Press: function_b14e0dd5("resetCounterUnlabel", 0)
   TextField "Text field_10" at 462,231 size 160x25; Text 'Labeled Counter'
   TextField "Text field_11" at 585,337 size 107x25; Text 'Label Time'
   TextField "Text field_12" at 123,213 size 108x25; Text 'Sorter Left'
   Circle "Circle_10" at 222,96 size 23x23
      Appearance <- "sorter"
   Circle "Circle_11" at 230,212 size 23x23
      Appearance <- "sorterLeft"
   TextField "Text field_5" at 129,355 size 102x25; Text 'Axis Label'
   Circle "Circle_12" at 236,354 size 23x23
      Appearance <- "axisLabel"
   TextField "Text field_22" at 674,229 size 158x25; Text 'Unlabel Counter'
   IOField "I/O field_2" at 567,378 size 136x56; FormatPattern 9
      ProcessValue <- "labelTime"
   TextField "Text field_8" at 1011,229 size 155x25; Text 'Sensors Signals'
   Circle "Circle_13" at 1002,303 size 23x23
      Appearance <- "heighBox"
   Circle "Circle_14" at 1002,333 size 23x23
      Appearance <- "positionBox"
   Circle "Circle_15" at 1002,363 size 23x23
      Appearance <- "unlabelBox"
   TextField "Text field_23" at 1059,299 size 102x25; Text 'Heigh Box'
   TextField "Text field_24" at 1059,332 size 125x25; Text 'Position Box'
   TextField "Text field_25" at 1058,362 size 119x25; Text 'Unlabel Box'
   Button "Button_1" at 82,140 size 97x47; TextOff 'Activate'
      on Press: InvertBit("activateSorter")
   Button "Button_2" at 200,140 size 97x47; TextOff 'Deactivate'
      on Press: InvertBit("activateSorter")
   Button "Button_3" at 82,271 size 97x47; TextOff 'Activate'
      on Press: InvertBit("activateSorterLeft")
   Button "Button_4" at 200,271 size 97x47; TextOff 'Deactivate'
      on Press: InvertBit("activateSorterLeft")
   Button "Button_5" at 82,402 size 97x47; TextOff 'Activate'
      on Press: InvertBit("activateAxis")
   Button "Button_6" at 200,402 size 97x47; TextOff 'Deactivate'
      on Press: InvertBit("activateAxis")
*)